   _43MB : ALIAS FOR B9[43].2;
   _43STB : ALIAS FOR B9[43].0;
   _43STPB : ALIAS FOR B9[43].1;
   _43Y : ALIAS FOR I25[2].14;
   _45_AIR_SEQ : ALIAS FOR T4[34];
   _45_AIR_SEQ1 : ALIAS FOR T4[34].PRE;
   _45_AIR_SEQ2 : ALIAS FOR T4[34].ACC;
   _45_SEQ_AIR : ALIAS FOR O12.15;
   _45AUTO : ALIAS FOR B9[45].4;
   _45HAND : ALIAS FOR B9[45].3;
   _45M : ALIAS FOR O25[8].7;
   _45MB : ALIAS FOR B9[45].2;
   _45STB : ALIAS FOR B9[45].0;
   _45STPB : ALIAS FOR B9[45].1;
   _45Y : ALIAS FOR I25[0].7;
   _46AUTO : ALIAS FOR B9[46].4;
   _46HAND : ALIAS FOR B9[46].3;
   _46M : ALIAS FOR O25[8].8;
   _46MB : ALIAS FOR B9[46].2;
   _46STB : ALIAS FOR B9[46].0;
   _46STPB : ALIAS FOR B9[46].1;
   _46Y : ALIAS FOR I25[0].8;
   _47AUTO : ALIAS FOR B9[47].4;
   _47HAND : ALIAS FOR B9[47].3;
   _47M : ALIAS FOR O25[9].10;
   _47MB : ALIAS FOR B9[47].2;
   _47STB : ALIAS FOR B9[47].0;
   _47STPB : ALIAS FOR B9[47].1;
   _47Y : ALIAS FOR I25[1].10;
   _48_CIMBRIA_HM : HOUR_METER := (MOTOR_RUNNING_INPUT_1 := 1, HR_METER_DISPLAY := 24757, MAINTENANCE_ALARM := 1);
   _48_FREQ_IN : ALIAS FOR N7[10];
   _48_FREQ_OU : ALIAS FOR N7[12];
   _48_SET_SPD : ALIAS FOR N7[11];
   _48_VFD_TO : ALIAS FOR N180[2];
   _48AUTO : ALIAS FOR B9[48].4;
   _48HAND : ALIAS FOR B9[48].3;
   _48M : ALIAS FOR O25[8].3;
   _48MAI : ALIAS FOR O25[25].2;
   _48MB : ALIAS FOR B9[48].2;
   _48STB : ALIAS FOR B9[48].0;
   _48STPB : ALIAS FOR B9[48].1;
   _48Y : ALIAS FOR I25[0].3;
   _49AUTO : ALIAS FOR B9[49].4;
   _49HAND : ALIAS FOR B9[49].3;
   _49M : ALIAS FOR O25[9].9;
   _49MB : ALIAS FOR B9[49].2;
   _49STB : ALIAS FOR B9[49].0;
   _49STPB : ALIAS FOR B9[49].1;
   _49Y : ALIAS FOR I25[1].9;
   _4_LOWER_TANK_CONVAYOR_21TO23_HM : HOUR_METER := (HR_METER_DISPLAY := 1470, NEXT_SCHDL_MAINTENANCE := 2, MAINTENANCE_ALARM := 1);
   _4_LOWER_TANK_CONVAYOR_21TO23_RUNNING : BOOL;
   _4_LS_TO_5 : ALIAS FOR I25[4].10;
   _4_LS_TO_6 : ALIAS FOR I25[4].11;
   _4_TO_BC5_S : ALIAS FOR O25[11].10;
   _4_TO_BC6_S : ALIAS FOR O25[11].11;
   _4AUTO : ALIAS FOR B9[4].4;
   _4HAND : ALIAS FOR B9[4].3;
   _4M : ALIAS FOR O25[10].1;
   _4MB : ALIAS FOR B9[4].2;
   _4STB : ALIAS FOR B9[4].0;
   _4STPB : ALIAS FOR B9[4].1;
   _4Y : ALIAS FOR I25[2].1;
   _50AUTO : ALIAS FOR B9[50].4;
   _50HAND : ALIAS FOR B9[50].3;
   _50M : ALIAS FOR O25[8].14;
   _50MB : ALIAS FOR B9[50].2;
   _50STB : ALIAS FOR B9[50].0;
   _50STPB : ALIAS FOR B9[50].1;
   _50Y : ALIAS FOR I25[0].14;
   _51_FREQ_IN : ALIAS FOR N7[13];
   _51_FREQ_OU : ALIAS FOR N7[15];
   _51_INDENT_HM : HOUR_METER := (MOTOR_RUNNING_INPUT_1 := 1, HR_METER_DISPLAY := 26515, MAINTENANCE_ALARM := 1);
   _51_SET_SPD : ALIAS FOR N7[14];
   _51_VFD_TO : ALIAS FOR N180[3];
   _51AUTO : ALIAS FOR B9[51].4;
   _51HAND : ALIAS FOR B9[51].3;
   _51M : ALIAS FOR O25[8].4;
   _51MAI : ALIAS FOR O25[25].3;
   _51MB : ALIAS FOR B9[51].2;
   _51STB : ALIAS FOR B9[51].0;
   _51STPB : ALIAS FOR B9[51].1;
   _51Y : ALIAS FOR I25[0].4;
   _52_FREQ_IN : ALIAS FOR N7[16];
   _52_FREQ_OU : ALIAS FOR N7[18];
   _52_SET_SPD : ALIAS FOR N7[17];
   _52AUTO : ALIAS FOR B9[52].4;
   _52HAND : ALIAS FOR B9[52].3;
   _52M : ALIAS FOR O25[8].6;
   _52MAI : ALIAS FOR O25[25].4;
   _52MB : ALIAS FOR B9[52].2;
   _52STB : ALIAS FOR B9[52].0;
   _52STPB : ALIAS FOR B9[52].1;
   _52Y : ALIAS FOR I25[0].6;
   _53_FREQ_IN : ALIAS FOR N7[7];
   _53_FREQ_OU : ALIAS FOR N7[9];
   _53_SET_SPD : ALIAS FOR N7[8];
   _53_VFD_TO : ALIAS FOR N180[1];
   _53AUTO : ALIAS FOR B9[53].4;
   _53HAND : ALIAS FOR B9[53].3;
   _53M : ALIAS FOR O25[8].2;
   _53MAI : ALIAS FOR O25[25].1;
   _53MB : ALIAS FOR B9[53].2;
   _53STB : ALIAS FOR B9[53].0;
   _53STPB : ALIAS FOR B9[53].1;
   _53Y : ALIAS FOR I25[0].2;
   _54AUTO : ALIAS FOR B9[54].4;
   _54HAND : ALIAS FOR B9[54].3;
   _54M : ALIAS FOR O25[11].3;
   _54MB : ALIAS FOR B9[54].2;
   _54STB : ALIAS FOR B9[54].0;
   _54STPB : ALIAS FOR B9[54].1;
   _54Y : ALIAS FOR I25[3].3;
   _55_FREQ_IN : ALIAS FOR N7[4];
   _55_FREQ_OU : ALIAS FOR N7[6];
   _55_SET_SPD : ALIAS FOR N7[5];
   _55AUTO : ALIAS FOR B9[55].4;
   _55HAND : ALIAS FOR B9[55].3;
   _55M : ALIAS FOR O25[8].1;
   _55MB : ALIAS FOR B9[55].2;
   _55STB : ALIAS FOR B9[55].0;
   _55STPB : ALIAS FOR B9[55].1;
   _55Y : ALIAS FOR I25[0].1;
   _56AUTO : ALIAS FOR B9[56].4;
   _56HAND : ALIAS FOR B9[56].3;
   _56M : ALIAS FOR O25[11].2;
   _56MB : ALIAS FOR B9[56].2;
   _56STB : ALIAS FOR B9[56].0;
   _56STPB : ALIAS FOR B9[56].1;
   _56Y : ALIAS FOR I25[3].2;
   _57AUTO : ALIAS FOR B9[57].4;
   _57HAND : ALIAS FOR B9[57].3;
   _57M : ALIAS FOR O25[9].6;
   _57MB : ALIAS FOR B9[57].2;
   _57STB : ALIAS FOR B9[57].0;
   _57STPB : ALIAS FOR B9[57].1;
   _57Y : ALIAS FOR I25[1].6;
   _5_LOWER_CROSS_BELT_HM : HOUR_METER := (HR_METER_DISPLAY := 2452, NEXT_SCHDL_MAINTENANCE := 2, MAINTENANCE_ALARM := 1);
   _5_LOWER_CROSS_BELT_RUNNING : BOOL;
   _5AUTO : ALIAS FOR B9[5].4;
   _5HAND : ALIAS FOR B9[5].3;
   _5M : ALIAS FOR O25[10].2;
   _5MB : ALIAS FOR B9[5].2;
   _5STB : ALIAS FOR B9[5].0;
   _5STPB : ALIAS FOR B9[5].1;
   _5Y : ALIAS FOR I25[2].2;
   _6AUTO : ALIAS FOR B9[6].4;
   _6HAND : ALIAS FOR B9[6].3;
   _6M : ALIAS FOR O25[10].3;
   _6MB : ALIAS FOR B9[6].2;
   _6STB : ALIAS FOR B9[6].0;
   _6STPB : ALIAS FOR B9[6].1;
   _6Y : ALIAS FOR I25[2].3;
   _700_AIR_GA : ALIAS FOR I8.3;
   _700_METER : ALIAS FOR I8.2;
   _700_PROBE : ALIAS FOR T22[9];
   _700_TREAT : ALIAS FOR I7.3;
   _700G_13_CL : ALIAS FOR B21[70].1;
   _700G_13_OP : ALIAS FOR B21[70].0;
   _700G_CLOSE : ALIAS FOR O12.9;
   _700G_OPEN : ALIAS FOR O12.8;
   _701_AIR_GA : ALIAS FOR I8.5;
   _701_FB : ALIAS FOR B21[1].3;
   _701_K_BYPA : ALIAS FOR I8.1;
   _701_K_TREA : ALIAS FOR I8.0;
   _701_METER : ALIAS FOR I8.4;
   _701_RB : ALIAS FOR B21[1].4;
   _701_REV_CN : ALIAS FOR C5[3];
   _701_STP : ALIAS FOR B21[1].2;
   _701_TRUCK_REVERSING_BELT_HM : HOUR_METER := (HR_METER_DISPLAY := 5981, NEXT_SCHDL_MAINTENANCE := 2, MAINTENANCE_ALARM := 1);
   _701_TRUCK_REVERSING_BELT_RUNNING : BOOL;
   _701F_HPB : ALIAS FOR B21[1].0;
   _701F_M : ALIAS FOR O25[10].11;
   _701F_OFF_T : ALIAS FOR T22[1];
   _701G_CLOSE : ALIAS FOR B21[71].13;
   _701G_OPEN : ALIAS FOR B21[71].12;
   _701K_GATE : ALIAS FOR B21[11].0;
   _701K_GATE1 : ALIAS FOR B21[11].1;
   _701K_GATE2 : ALIAS FOR B21[11].2;
   _701K_VALVE : ALIAS FOR O13.10;
   _701MR : ALIAS FOR O25[9].7;
   _701R_DELAY : ALIAS FOR T22[2];
   _701R_HPB : ALIAS FOR B21[1].1;
   _701Y : BOOL;
   _701YF : ALIAS FOR I25[2].11;
   _701YR : ALIAS FOR I25[1].7;
   _702_CLEAN_JUMP_BELT_HM : HOUR_METER := (HR_METER_DISPLAY := 3983, NEXT_SCHDL_MAINTENANCE := 2, MAINTENANCE_ALARM := 1);
   _702B : ALIAS FOR B21[2].2;
   _702H_START : ALIAS FOR B21[2].0;
   _702H_STOP : ALIAS FOR B21[2].1;
   _702M : ALIAS FOR O25[9].4;
   _702Y : ALIAS FOR I25[1].4;
   _703_TREATER_JUMP_BELT_HM : HOUR_METER := (HR_METER_DISPLAY := 2423, NEXT_SCHDL_MAINTENANCE := 2, MAINTENANCE_ALARM := 1);
   _703_TREATER_JUMP_BELT_RUNNING : BOOL;
   _703B : ALIAS FOR B21[3].2;
   _703H_START : ALIAS FOR B21[3].0;
   _703H_STOP : ALIAS FOR B21[3].1;
   _703M : ALIAS FOR O25[9].14;
   _703Y : ALIAS FOR I25[1].14;
   _704B : ALIAS FOR B21[4].2;
   _704H_START : ALIAS FOR B21[4].0;
   _704H_STOP : ALIAS FOR B21[4].1;
   _704M : ALIAS FOR O25[8].11;
   _704Y : ALIAS FOR I25[0].13;
   _705B : ALIAS FOR B21[5].2;
   _705H_START : ALIAS FOR B21[5].0;
   _705H_STOP : ALIAS FOR B21[5].1;
   _705M : ALIAS FOR O25[10].12;
   _705Y : ALIAS FOR I25[2].12;
   _705YA : ALIAS FOR I25[4].15;
   _706B : ALIAS FOR B21[6].2;
   _706H_START : ALIAS FOR B21[6].0;
   _706H_STOP : ALIAS FOR B21[6].1;
   _706M : ALIAS FOR O25[9].11;
   _706Y : ALIAS FOR I25[1].11;
   _707B : ALIAS FOR B21[7].2;
   _707M : ALIAS FOR O25[11].0;
   _707Y : ALIAS FOR I25[3].0;
   _708_BOT_CN : ALIAS FOR C5[5];
   _708G_BIN_1 : ALIAS FOR O9.15;
   _708G_BIN_2 : ALIAS FOR I7.4;
   _708G_CB13 : ALIAS FOR B21[8].0;
   _708G_CB131 : ALIAS FOR B21[8].1;
   _708G_CB132 : ALIAS FOR B21[8].2;
   _708G_HOLD : ALIAS FOR B21[8].3;
   _708G_HOLD1 : ALIAS FOR B21[8].6;
   _708G_RELEA : ALIAS FOR B21[8].4;
   _708G_RESET : ALIAS FOR B21[8].5;
   _709_BOT_CN : ALIAS FOR C5[6];
   _709G_BIN_1 : ALIAS FOR O10.15;
   _709G_BIN_2 : ALIAS FOR I7.5;
   _709G_CB19 : ALIAS FOR B21[9].0;
   _709G_CB191 : ALIAS FOR B21[9].1;
   _709G_CB192 : ALIAS FOR B21[9].2;
   _709G_HOLD : ALIAS FOR B21[9].3;
   _709G_HOLD1 : ALIAS FOR B21[9].6;
   _709G_RELEA : ALIAS FOR B21[9].4;
   _709G_RESET : ALIAS FOR B21[9].5;
   _709G_RUN_T : ALIAS FOR T22[8];
   _709G_TREAT : ALIAS FOR B21[9].7;
   _709G_TREAT1 : ALIAS FOR T22[10];
   _7AUTO : ALIAS FOR B9[7].4;
   _7HAND : ALIAS FOR B9[7].3;
   _7MB : ALIAS FOR B9[7].2;
   _7STB : ALIAS FOR B9[7].0;
   _7STPB : ALIAS FOR B9[7].1;
   _8AUTO : ALIAS FOR B9[8].4;
   _8HAND : ALIAS FOR B9[8].3;
   _8MB : ALIAS FOR B9[8].2;
   _8STB : ALIAS FOR B9[8].0;
   _8STPB : ALIAS FOR B9[8].1;
   _9_AIR_SV : ALIAS FOR O24[7].6;
   _9_BYPSS_GT : ALIAS FOR I24[6].1;
   _9_CAL_MOV : ALIAS FOR O24[7].2;
   _9_CAL_VALV : ALIAS FOR I24[6].5;
   _9_DRIP_GAT : ALIAS FOR O24[7].7;
   _9_GATE_SV : ALIAS FOR O24[7].0;
   _9_GATE_SV1 : ALIAS FOR O24[7].1;
   _9_SL_SW : ALIAS FOR B9[9].6;
   _9_SLW_SPEE : ALIAS FOR I25[3].12;
   _9_STP_SPEE : ALIAS FOR I25[3].13;
   _9_TREAT_MV : ALIAS FOR I24[6].6;
   _9_TREATER : ALIAS FOR I24[6].7;
   _9_TREATER_CONVAYOR_HM : HOUR_METER := (HR_METER_DISPLAY := 4578, NEXT_SCHDL_MAINTENANCE := 2, MAINTENANCE_ALARM := 1);
   _9_TREATER_CONVAYOR_RUNNING : BOOL;
   _9_TRT_M_ST : ALIAS FOR I24[6].3;
   _9_TRT_M_ST1 : ALIAS FOR I24[6].4;
   _9_TRT_MB : ALIAS FOR B3[9].0;
   _9_TRT_MOV : ALIAS FOR O24[7].4;
   _9_TRT_STB : ALIAS FOR B3[9].1;
   _9_TRT_STPB : ALIAS FOR B3[9].2;
   _9AUTO : ALIAS FOR B9[9].4;
   _9HAND : ALIAS FOR B9[9].3;
   _9M : ALIAS FOR O25[8].10;
   _9MB : ALIAS FOR B9[9].2;
   _9STB : ALIAS FOR B9[9].0;
   _9STPB : ALIAS FOR B9[9].1;
   _9Y : ALIAS FOR I25[0].10;
   _9YB : ALIAS FOR B9[9].5;
   A16 : INT[250] := ([24] := '0 ', [25] := '0 ', [26] := '0 ', [48] := '0 ', [110] := 'ge', [140] := 'ha', [150] := '10', [200] := 'cl', [210] := 'ov', [240] := 'le');
   A18 : INT[100] := ([13] := '9$00');
   A_ACC : ALIAS FOR N10[11];
   A_ACC_SEC : ALIAS FOR N10[13];
   A_HOLD_B : ALIAS FOR B3[1].4;
   A_HOLD_MB : ALIAS FOR B3[1].3;
   A_HOLD_REL : ALIAS FOR B3[1].5;
   A_MAIN_CNT : ALIAS FOR C5[0].PRE;
   A_MAIN_CNT1 : ALIAS FOR C5[0].ACC;
   A_MAIN_TRE : ALIAS FOR C5[0];
   A_PRESET : ALIAS FOR N10[10];
   A_PRESET_S : ALIAS FOR N10[12];
   A_RESET_PB : ALIAS FOR B3[1].2;
   A_SET : ALIAS FOR B3[1].6;
   A_STB_AUTO : ALIAS FOR B3[1].0;
   A_STPB_AUT : ALIAS FOR B3[1].1;
   A_TREATER : ALIAS FOR I24[6].8;
   A_TREATER1 : ALIAS FOR T4[59];
   ALARM_FIEL : ALIAS FOR T11[7];
   ALARM_HAND : ALIAS FOR B3[0].10;
   ALARM_HMI : ALIAS FOR B3[0].6;
   ALARM_HORN : ALIAS FOR O25[11].15;
   ALARM_HORN1 : ALIAS FOR O12.14;
   ALARM_INIT : ALIAS FOR B3[0].4;
   ALARM_LIGH : ALIAS FOR O13.15;
   ALARM_LT_O : ALIAS FOR T11[3];
   ALARM_SILE : ALIAS FOR I25[4].7;
   ALARM_SILE1 : ALIAS FOR I7.13;
   ALARM_SILE2 : ALIAS FOR B3[0].3;
   ALARM_SILE3 : ALIAS FOR B3[0].5;
   ALARM_SILE4 : ALIAS FOR B3[0].9;
   ALRM_LIGHT : ALIAS FOR O25[11].14;
   ALRM_SILEN : ALIAS FOR B3[0].7;
   Always_On : BOOL := 1;
   Analog : AI[160] := ([0].In := 104.0, [0].RawMin := 147.0, [0].RawMax := 16384.0, [0].EUMax := 3770.0, [1].In := 131.0, [1].RawMin := 147.0, [1].RawMax := 16384.0, [1].EUMax := 3770.0, [2].In := 1848.0, [2].RawMin := 1884.0, [2].RawMax := 16384.0, [2].EUMax := 4000.0, [20].In := 28816.0, [20].RawMin := 31000.0, [20].EUMax := 3200.0, [20].Out := 2974.5547, [21].In := 30336.0, [21].RawMax := 31000.0, [21].EUMax := 3200.0, [21].Out := 3131.458, [22].In := 30064.0, [22].RawMax := 31000.0, [22].EUMax := 3200.0, [22].Out := 3103.3806, [23].In := 7360.0, [23].RawMax := 31000.0, [23].EUMax := 3200.0, [23].Out := 759.74194, [24].In := 9136.0, [24].RawMax := 31000.0, [24].EUMax := 3200.0, [24].Out := 943.0709, [25].In := 28656.0, [25].RawMax := 31000.0, [25].EUMax := 3200.0, [25].Out := 2958.0386, [26].In := 28944.0, [26].RawMax := 31000.0, [26].EUMax := 3200.0, [26].Out := 2987.7676);
   B12 : DINT[100];
   B15 : DINT[100] := ([16] := 2#0000_0000_0000_0000_0000_0000_0000_0011, [17] := 2#0000_0000_0000_0000_0000_0000_0000_0011, [21] := 2#0000_0000_0000_0000_0000_0000_0000_0011, [22] := 2#0000_0000_0000_0000_0000_0000_0000_0011, [23] := 2#0000_0000_0000_0000_0000_0000_0000_0011, [30] := 2#0000_0000_0000_0000_0000_0000_0000_0011);
   B17 : DINT[30] := ([11] := 2#0000_0000_0000_0000_0000_0000_0000_0010, [12] := 2#0000_0000_0000_0000_0000_0000_0000_0111, [13] := 2#0000_0000_0000_0000_0000_0000_0000_0111, [14] := 2#0000_0000_0000_0000_0000_0000_0000_0010, [15] := 2#0000_0000_0000_0000_0000_0000_0000_0010, [16] := 2#0000_0000_0000_0000_0000_0000_0000_0111, [17] := 2#0000_0000_0000_0000_0000_0000_0000_0111, [21] := 2#0000_0000_0000_0000_0000_0000_0000_0010, [22] := 2#0000_0000_0000_0000_0000_0000_0000_0111, [23] := 2#0000_0000_0000_0000_0000_0000_0000_0111, [24] := 2#0000_0000_0000_0000_0000_0000_0000_0010, [25] := 2#0000_0000_0000_0000_0000_0000_0000_0111, [26] := 2#0000_0000_0000_0000_0000_0000_0000_0010);
   B183 : DINT[1] := ([0] := 2#0000_0000_0000_0000_0000_0000_0000_0001);
   B184 : DINT[1] := ([0] := 2#0000_0000_0000_0000_0000_0000_0000_0010);
   B194 : DINT[1];
   B204 : DINT[1];
   B21 : DINT[255];
   B214 : DINT[1];
   B224 : DINT[1] := ([0] := 2#0000_0000_0000_0000_0000_0000_0000_0010);
   B234 : DINT[1];
   B243 : DINT[1] := ([0] := 2#0000_0000_0000_0000_0000_0000_0000_0011);
   B244 : DINT[1] := ([0] := 2#0000_0000_0000_0000_0000_0000_0000_0010);
   B253 : DINT[100] := ([0] := 2#0000_0000_0000_0000_0000_0000_0000_0011);
   B254 : DINT[1] := ([0] := 2#0000_0000_0000_0000_0000_0000_0000_0010);
   B3 : DINT[250] := ([0] := 2#0000_0000_0000_0000_0000_0010_1011_0000, [101] := 2#0000_0000_0000_0000_0000_0000_0000_0010, [102] := 2#0000_0000_0000_0000_0000_0000_1000_0001);
   B9 : DINT[150] := ([1] := 2#0000_0000_0000_0000_0000_0000_0001_0100, [35] := 2#0000_0000_0000_0000_0000_0000_0001_0100, [42] := 2#0000_0000_0000_0000_0000_0000_0001_0100, [43] := 2#0000_0000_0000_0000_0000_0000_0011_0100, [45] := 2#0000_0000_0000_0000_0000_0000_0001_0100, [46] := 2#0000_0000_0000_0000_0000_0000_0001_0100, [48] := 2#0000_0000_0000_0000_0000_0000_0001_0100, [49] := 2#0000_0000_0000_0000_0000_0000_0001_0100, [50] := 2#0000_0000_0000_0000_0000_0000_0000_1000, [51] := 2#0000_0000_0000_0000_0000_0000_0001_0100, [52] := 2#0000_0000_0000_0000_0000_0000_0001_0100, [53] := 2#0000_0000_0000_0000_0000_0000_0001_0100, [54] := 2#0000_0000_0000_0000_0000_0000_0001_0100, [55] := 2#0000_0000_0000_0000_0000_0000_0001_0100, [57] := 2#0000_0000_0000_0000_0000_0000_0001_0100, [102] := 2#0000_0000_0000_0000_0000_0000_0000_1000, [103] := 2#0000_0000_0000_0000_0000_0000_0000_1000, [107] := 2#0000_0000_0000_0000_0000_0000_0011_0100, [108] := 2#0000_0000_0000_0000_0000_0000_0001_0100, [122] := 2#0000_0000_0000_0000_0000_0000_0001_0100, [123] := 2#0000_0000_0000_0000_0000_0000_0001_0100);
   Beta : BOOL := 1;
   BIN_1_CLOSE : BOOL;
   BIN_1_OPEN : BOOL;
   BIN_2_CLOSE : BOOL;
   BIN_2_OPEN : BOOL;
   BIN_3_CLOSE : BOOL;
   BIN_3_OPEN : BOOL;
   BIN_4_CLOSE : BOOL;
   BIN_4_OPEN : BOOL;
   BIN_5_CLOSE : BOOL;
   BIN_5_OPEN : BOOL;
   BIN_6_CLOSE : BOOL;
   BIN_6_OPEN : BOOL;
   BIN_7_CLOSE : BOOL;
   BIN_7_OPEN : BOOL;
   Bin_Config : BOOL := 1;
   C5 : COUNTER[50] := ([0].PRE := 3000, [1].ACC := 5, [1].DN := 1, [2].PRE := 3000, [3].PRE := 2, [4].PRE := 400000, [5].PRE := 5000, [5].CU := 1, [6].PRE := 9999, [6].CU := 1, [11].PRE := 1200, [12].PRE := 30, [13].PRE := 3000, [14].PRE := 36, [15].PRE := 1500, [16].PRE := 3000, [17].PRE := 3000, [21].PRE := 3000, [22].PRE := 3000, [23].PRE := 3000, [24].PRE := 3000, [25].PRE := 3000, [26].PRE := 3000, [27].CU := 1, [28].CU := 1, [29].CU := 1, [30].PRE := 20000, [32].PRE := 20000, [33].PRE := 20000, [34].PRE := 20000, [35].PRE := 20000, [36].PRE := 20000, [37].PRE := 20000, [38].PRE := 20000, [39].PRE := 20000);
   CAL_K_FACT : ALIAS FOR F8[0];
   CAL_RESET : ALIAS FOR B15[50].0;
   Calibration_Max : REAL := 4000.0;
   CG13_METR : ALIAS FOR I8.15;
   CG_13_AIR : ALIAS FOR I8.13;
   CG_19_AIR : ALIAS FOR I8.12;
   CG_19_METR : ALIAS FOR I8.14;
   CHEM_PUMP_1 : STRING := 'water';
   CHEM_PUMP_10 : STRING := 'oil';
   CHEM_PUMP_11 : STRING := 'apron';
   CHEM_PUMP_12 : STRING := 'stamina';
   CHEM_PUMP_13 : STRING := 'TEST13';
   CHEM_PUMP_14 : STRING := 'oil';
   CHEM_PUMP_15 : STRING := 'red';
   CHEM_PUMP_2 : STRING := 'alba red';
   CHEM_PUMP_3 : STRING := 'evergol';
   CHEM_PUMP_4 : STRING := 'macho';
   CHEM_PUMP_5 : STRING := 'vib ex';
   CHEM_PUMP_6 : STRING := 'bio st';
   CHEM_PUMP_7 : STRING := 'tbz';
   CHEM_PUMP_8 : STRING := 'wuxal';
   CHEM_PUMP_9 : STRING := 'BLUE';
   CIMBRA_BIN : ALIAS FOR I25[3].10;
   CIMBRIA_BI : ALIAS FOR B15[30].0;
   CIMBRIA_BI1 : ALIAS FOR B15[30].1;
   CIMBRIA_BIN_EMPTY : BOOL;
   CIMBRIA_BIN_FULL : BOOL;
   CIMBRIA_FAN_ON : BOOL := 1;
   CIMBRIA_FAN_SPD_INPUT : DINT := 30;
   CIMBRIA_HI : ALIAS FOR B15[30].2;
   CIMBRIA_OUTPUT_SPD : DINT := 30;
   Cleaning_Motors : udt_Motor[100] := ([0].Motor_Control.Motor_Amps := 1.3896561, [1].Motor_Control.Motor_Amps := 1.006918, [2].Motor_Control.Motor_Amps := 0.8792738, [3].Motor_Control.Motor_Amps := 2.5666564);
   CLR_SORT_ASP_DELAY : TIMER := (PRE := 5000, ACC := 5002, EN := 1, DN := 1);
   CLR_SORT_ASPBLR_DELAY : TIMER := (PRE := 5000, ACC := 5004, EN := 1, DN := 1);
   CLR_SORT_LEG_DELAY : TIMER := (PRE := 5000, ACC := 5003, EN := 1, DN := 1);
   CLR_SORT_LEG_SPD10 : ALIAS FOR Local:0:I.Data.3;
   CLR_SORT_LEG_SPD20 : ALIAS FOR Local:0:I.Data.4;
   CONC13_COL : ALIAS FOR N7[93];
   CONC13_OP : ALIAS FOR A18[3];
   CONC13_PUM : ALIAS FOR N7[83];
   CONC13_SET : ALIAS FOR A18[0];
   CONC13_SET1 : ALIAS FOR B21[8].14;
   CONC19_COL : ALIAS FOR N7[99];
   CONC19_OP : ALIAS FOR A18[13];
   CONC19_PUM : ALIAS FOR N7[89];
   CONC19_SET : ALIAS FOR B21[9].14;
   CONC_13_NO : ALIAS FOR B21[8].15;
   CONC_19_NO : ALIAS FOR B21[9].15;
   CONC_19_SE : ALIAS FOR A18[10];
   ConcretePlantIn : DINT := 2;
   ConcretePlantOut : DINT := 1; {produced}
   Config_Save_Binss : BOOL;
   ConfigureVariety : Variety;
   Consumed : DINT;
   CP_Remote_Air_Gate_On : DINT; {produced}
   CP_Remote_Air_Gate_Open_In : DINT;
   CP_Remote_Andco_Auto_In : DINT;
   CP_Remote_Andoc_Out : udt_Andco_Remote_Out[32]; {produced}
   CP_Remote_Belt_In : udt_Motor_Remote_In[10] := ([1].Spd_10_Out := 1, [1].Amps := -0.32500002, [2].Spd_10_Out := 1, [2].Amps := -0.425, [3].Spd_10_Out := 1, [3].Amps := -0.5125);
   CP_Remote_Belt_Start : DINT; {produced}
   CP_Remote_Leg_In : udt_Motor_Remote_In := (Spd_20_Out := 1, Spd_10_Out := 1, Amps := -0.22500001);
   CP_Remote_Leg_Start : DINT; {produced}
   cpBinGateRates : DINT[50] := ([1] := 73, [3] := 180, [5] := 531, [7] := 117, [10] := 147, [13] := 269, [19] := 173);
   cpBINOPEN : DINT;
   cpCleanBulk : BOOL;
   cpTicketBinActive : DINT;
   cpTicketBinSet : DINT;
   cpVAR_BINARRAY : STRING[50] := ([1] := '823019-Diva Spring-Certified-WSU -SWW Seed Wheat', [3] := '823007-WB 6121 spring-Certified - Monsanto  - SWW Seed Wheat', [4] := 'reg duet', [5] := '823001-ArtDeco-Certified-Limagrain -SWW Seed Wheat', [10] := '823007-WB 6121 spring-Certified-Monsanto -SWW Seed Wheat', [11] := '823014-Skiles-Certified-OSU -SWW Seed Wheat', [20] := '823010-Bobtail-Certified-OSU -SWW Seed Wheat');
   cpVAR_CNT_ONS : DINT;
   cpVarTrimTemp : STRING := '823026';
   Dev : DINT := 6145; {produced}
   DIST_MOVE : ALIAS FOR I3.10;
   DIST_TO_CL : ALIAS FOR I7.2;
   DS_CLEAN_B : ALIAS FOR O13.5;
   DS_DLY_OFF : ALIAS FOR T4[33];
   DS_M : ALIAS FOR O24[1].0;
   DS_M_B : ALIAS FOR B3[101].0;
   DS_MOV_CCW : ALIAS FOR B3[100].13;
   DS_MOV_CW : ALIAS FOR B3[100].12;
   DS_MOVE_SE : ALIAS FOR T4[32];
   DS_POS8 : ALIAS FOR O13.7;
   DS_POS9 : ALIAS FOR O13.8;
   DS_POS_1 : ALIAS FOR I24[0].2;
   DS_POS_10 : ALIAS FOR I24[0].11;
   DS_POS_11 : ALIAS FOR B3[100].11;
   DS_POS_1_B : ALIAS FOR B3[100].2;
   DS_POS_2 : ALIAS FOR I24[0].3;
   DS_POS_2_B : ALIAS FOR B3[100].3;
   DS_POS_3 : ALIAS FOR I24[0].4;
   DS_POS_3_B : ALIAS FOR B3[100].4;
   DS_POS_4 : ALIAS FOR I24[0].5;
   DS_POS_4_B : ALIAS FOR B3[100].5;
   DS_POS_5 : ALIAS FOR I24[0].6;
   DS_POS_5_B : ALIAS FOR B3[100].6;
   DS_POS_6 : ALIAS FOR I24[0].7;
   DS_POS_6_B : ALIAS FOR B3[100].7;
   DS_POS_7 : ALIAS FOR I24[0].8;
   DS_POS_7_B : ALIAS FOR B3[100].8;
   DS_POS_8 : ALIAS FOR I24[0].9;
   DS_POS_8_B : ALIAS FOR B3[100].9;
   DS_POS_9 : ALIAS FOR I24[0].10;
   DS_POS_9_B : ALIAS FOR B3[100].10;
   DS_SEEK_1 : ALIAS FOR B3[102].1;
   DS_SEEK_10 : ALIAS FOR B3[102].10;
   DS_SEEK_2 : ALIAS FOR B3[102].2;
   DS_SEEK_3 : ALIAS FOR B3[102].3;
   DS_SEEK_4 : ALIAS FOR B3[102].4;
   DS_SEEK_5 : ALIAS FOR B3[102].5;
   DS_SEEK_6 : ALIAS FOR B3[102].6;
   DS_SEEK_7 : ALIAS FOR B3[102].7;
   DS_SEEK_8 : ALIAS FOR B3[102].8;
   DS_SEEK_9 : ALIAS FOR B3[102].9;
   DS_SET_IN : ALIAS FOR N10[0];
   DS_SP_UP_B : ALIAS FOR B3[100].0;
   DS_SPOUT_C : ALIAS FOR O24[1].3;
   DS_SPOUT_C1 : ALIAS FOR O24[1].4;
   DS_SPOUT_C2 : ALIAS FOR B3[101].3;
   DS_SPOUT_C3 : ALIAS FOR B3[101].4;
   DS_SPOUT_D : ALIAS FOR I24[0].1;
   DS_SPOUT_D1 : ALIAS FOR O24[1].1;
   DS_SPOUT_D2 : ALIAS FOR B3[100].1;
   DS_SPOUT_D3 : ALIAS FOR B3[101].1;
   DS_SPOUT_U : ALIAS FOR I24[0].0;
   DS_SPOUT_U1 : ALIAS FOR O24[1].2;
   DS_SPOUT_U2 : ALIAS FOR B3[101].2;
   DS_START_M : ALIAS FOR B3[102].11;
   DS_STOP_MO : ALIAS FOR B3[102].0;
   DS_T21 : ALIAS FOR O13.0;
   DS_T22 : ALIAS FOR O13.1;
   DS_T23 : ALIAS FOR O13.9;
   DS_T231 : ALIAS FOR O13.2;
   DS_T24 : ALIAS FOR O13.3;
   DS_T25 : ALIAS FOR O13.4;
   DS_T26 : ALIAS FOR O13.6;
   F8 : REAL[27] := ([0] := 1.2, [1] := 1.0, [2] := 14748.0, [3] := 1.0, [4] := 15440.0, [5] := 1.0, [6] := 14244.0, [7] := 1.0, [8] := 13454.0, [9] := 1.0, [10] := 14460.0, [11] := 1.0, [12] := 6343.0, [13] := 1.0, [14] := 8758.0, [15] := 1.0, [16] := 15944.0, [17] := 1.0, [18] := 15184.0, [19] := 1.0, [20] := 15741.0, [21] := 1.0, [22] := 15276.0, [23] := 1.0, [24] := 14611.0, [25] := 1.0, [26] := 15145.0);
   Gates : STRING;
   hCLR_SORT_LEG_SPD10 : BOOL := 1;
   hCLR_SORT_LEG_SPD20 : BOOL := 1;
   hCLR_SORT_STB : BOOL;
   hCLR_SORT_STRT : BOOL;
   hN_RECVING_PIT_GATE_CLSPB : BOOL;
   hN_RECVING_PIT_GATE_OPNPB : BOOL;
   hSURGE_BIN_HI : BOOL;
   hSURGE_BIN_LO : BOOL;
   I1 : ALIAS FOR R1S0_AENTR:1:I.Data;
   I16 : INT[16] := ([0] := 2#0011_1001_1001_1100, [1] := 2#0011_1100_0101_0000, [2] := 2#0011_0111_1010_0100, [3] := 2#0011_0100_1000_1110, [4] := 2#0011_1000_0111_1100, [5] := 2#0001_1000_1100_0111, [6] := 2#0010_0010_0011_0110, [7] := 2#0011_1110_0100_1000, [8] := 2#0000_1000_0101_1010, [9] := 2#0000_1000_0101_1010, [10] := 2#0000_1000_0101_1010, [11] := 2#0000_1000_0101_1010, [12] := 2#0000_1000_0101_1010, [13] := 2#0000_1000_0101_1010, [14] := 2#0000_1000_0101_1010, [15] := 2#0000_1000_0101_1010);
   I16_0 : ALIAS FOR N20[0];
   I16_000 : ALIAS FOR I16[0];
   I16_001 : ALIAS FOR I16[1];
   I16_002 : ALIAS FOR I16[2];
   I16_003 : ALIAS FOR I16[3];
   I16_004 : ALIAS FOR I16[4];
   I16_005 : ALIAS FOR I16[5];
   I16_006 : ALIAS FOR I16[6];
   I16_007 : ALIAS FOR I16[7];
   I16_1 : ALIAS FOR N20[1];
   I16_2 : ALIAS FOR N20[2];
   I16_3 : ALIAS FOR N20[3];
   I16_4 : ALIAS FOR N20[4];
   I16_5 : ALIAS FOR N20[5];
   I16_6 : ALIAS FOR N20[6];
   I16_7 : ALIAS FOR N20[7];
   I17 : INT[16] := ([0] := 2#0011_1011_0101_0000, [1] := 2#0011_1101_0111_1101, [2] := 2#0011_1011_1010_1111, [3] := 2#0011_1001_0001_0011, [4] := 2#0011_1011_0010_1001, [5] := 2#0001_1100_1010_0101, [6] := 2#0001_1100_1010_1111, [7] := 2#0001_1100_1010_0010, [8] := 2#0000_1000_0101_1010, [9] := 2#0000_1000_0101_1010, [10] := 2#0000_1000_0101_1010, [11] := 2#0000_1000_0101_1010, [12] := 2#0000_1000_0101_1010, [13] := 2#0000_1000_0101_1010, [14] := 2#0000_1000_0101_1010, [15] := 2#0000_1000_0101_1010);
   I17_000 : ALIAS FOR I17[0];
   I17_001 : ALIAS FOR I17[1];
   I17_002 : ALIAS FOR I17[2];
   I17_003 : ALIAS FOR I17[3];
   I17_004 : ALIAS FOR I17[4];
   I17_005 : ALIAS FOR I17[5];
   I17_006 : ALIAS FOR I17[6];
   I17_007 : ALIAS FOR I17[7];
   I18 : INT[16] := ([0] := 2#0000_0101_0101_0011, [1] := 2#0000_0111_0011_1000, [2] := 2#0000_0000_1000_0011, [3] := 2#0000_0000_0110_1000, [4] := 2#0000_0111_0111_1100, [5] := 2#0000_0111_0110_0101, [6] := 2#0000_1100_1100_1101, [7] := 2#0000_1100_1100_1101, [8] := 2#0000_1000_0101_1010, [9] := 2#0000_1000_0101_1010, [10] := 2#0000_1000_0101_1010, [11] := 2#0000_1000_0101_1010, [12] := 2#0000_1000_0101_1010, [13] := 2#0000_1000_0101_1010, [14] := 2#0001_1010_1001_1101, [15] := 2#0001_1010_1001_1101);
   I18_000 : ALIAS FOR I18[0];
   I18_001 : ALIAS FOR I18[1];
   I18_002 : ALIAS FOR I18[2];
   I18_003 : ALIAS FOR I18[3];
   I18_007 : ALIAS FOR I18[7];
   I1_000_Bit00 : ALIAS FOR I1.0;
   I1_000_Bit01 : ALIAS FOR I1.1;
   I1_000_Bit02 : ALIAS FOR I1.2;
   I1_000_Bit03 : ALIAS FOR I1.3;
   I1_000_Bit04 : ALIAS FOR I1.4;
   I1_000_Bit05 : ALIAS FOR I1.5;
   I1_000_Bit06 : ALIAS FOR I1.6;
   I1_000_Bit07 : ALIAS FOR I1.7;
   I1_000_Bit08 : ALIAS FOR I1.8;
   I1_000_Bit09 : ALIAS FOR I1.9;
   I1_000_Bit10 : ALIAS FOR I1.10;
   I1_000_Bit11 : ALIAS FOR I1.11;
   I1_000_Bit12 : ALIAS FOR I1.12;
   I1_000_Bit13 : ALIAS FOR I1.13;
   I1_000_Bit14 : ALIAS FOR I1.14;
   I1_000_Bit15 : ALIAS FOR I1.15;
   I2 : ALIAS FOR R1S0_AENTR:2:I.Data;
   I24 : INT[32] := ([0] := 2#0000_0001_0000_0010, [6] := 2#0010_0000_1000_0110, [7] := 2#0010_0000_1000_0110);
   I24_000_Bit00 : ALIAS FOR I24[0].0;
   I24_000_Bit01 : ALIAS FOR I24[0].1;
   I24_000_Bit02 : ALIAS FOR I24[0].2;
   I24_000_Bit03 : ALIAS FOR I24[0].3;
   I24_000_Bit04 : ALIAS FOR I24[0].4;
   I24_000_Bit05 : ALIAS FOR I24[0].5;
   I24_000_Bit06 : ALIAS FOR I24[0].6;
   I24_000_Bit07 : ALIAS FOR I24[0].7;
   I24_000_Bit08 : ALIAS FOR I24[0].8;
   I24_000_Bit09 : ALIAS FOR I24[0].9;
   I24_000_Bit10 : ALIAS FOR I24[0].10;
   I24_000_Bit11 : ALIAS FOR I24[0].11;
   I24_004_Bit00 : ALIAS FOR I24[4].0;
   I24_004_Bit01 : ALIAS FOR I24[4].1;
   I24_004_Bit02 : ALIAS FOR I24[4].2;
   I24_004_Bit03 : ALIAS FOR I24[4].3;
   I24_004_Bit04 : ALIAS FOR I24[4].4;
   I24_004_Bit05 : ALIAS FOR I24[4].5;
   I24_004_Bit06 : ALIAS FOR I24[4].6;
   I24_004_Bit07 : ALIAS FOR I24[4].7;
   I24_004_Bit08 : ALIAS FOR I24[4].8;
   I24_004_Bit09 : ALIAS FOR I24[4].9;
   I24_004_Bit10 : ALIAS FOR I24[4].10;
   I24_004_Bit11 : ALIAS FOR I24[4].11;
   I24_004_Bit12 : ALIAS FOR I24[4].12;
   I24_006_Bit01 : ALIAS FOR I24[6].1;
   I24_006_Bit02 : ALIAS FOR I24[6].2;
   I24_006_Bit07 : ALIAS FOR I24[6].7;
   I24_006_Bit08 : ALIAS FOR I24[6].8;
   I24_006_Bit13 : ALIAS FOR I24[6].13;
   I24_021_Bit00 : ALIAS FOR I24[21].0;
   I24_021_Bit01 : ALIAS FOR I24[21].1;
   I24_021_Bit02 : ALIAS FOR I24[21].2;
   I24_021_Bit03 : ALIAS FOR I24[21].3;
   I24_021_Bit04 : ALIAS FOR I24[21].4;
   I24_021_Bit05 : ALIAS FOR I24[21].5;
   I24_021_Bit06 : ALIAS FOR I24[21].6;
   I24_021_Bit07 : ALIAS FOR I24[21].7;
   I24_021_Bit08 : ALIAS FOR I24[21].8;
   I25 : INT[32] := ([0] := 2#0101_0011_1101_1110, [1] := 2#0011_0011_0100_0010, [2] := 2#1110_0000_0100_0000, [3] := 2#1101_0000_0000_1010, [4] := 2#0110_0000_0000_1101);
   I25_000_Bit00 : ALIAS FOR I25[0].0;
   I25_000_Bit01 : ALIAS FOR I25[0].1;
   I25_000_Bit02 : ALIAS FOR I25[0].2;
   I25_000_Bit03 : ALIAS FOR I25[0].3;
   I25_000_Bit04 : ALIAS FOR I25[0].4;
   I25_000_Bit06 : ALIAS FOR I25[0].6;
   I25_000_Bit07 : ALIAS FOR I25[0].7;
   I25_000_Bit08 : ALIAS FOR I25[0].8;
   I25_000_Bit09 : ALIAS FOR I25[0].9;
   I25_000_Bit10 : ALIAS FOR I25[0].10;
   I25_000_Bit12 : ALIAS FOR I25[0].12;
   I25_000_Bit13 : ALIAS FOR I25[0].13;
   I25_000_Bit14 : ALIAS FOR I25[0].14;
   I25_000_Bit15 : ALIAS FOR I25[0].15;
   I25_001_Bit00 : ALIAS FOR I25[1].0;
   I25_001_Bit01 : ALIAS FOR I25[1].1;
   I25_001_Bit02 : ALIAS FOR I25[1].2;
   I25_001_Bit03 : ALIAS FOR I25[1].3;
   I25_001_Bit04 : ALIAS FOR I25[1].4;
   I25_001_Bit05 : ALIAS FOR I25[1].5;
   I25_001_Bit06 : ALIAS FOR I25[1].6;
   I25_001_Bit07 : ALIAS FOR I25[1].7;
   I25_001_Bit08 : ALIAS FOR I25[1].8;
   I25_001_Bit09 : ALIAS FOR I25[1].9;
   I25_001_Bit10 : ALIAS FOR I25[1].10;
   I25_001_Bit11 : ALIAS FOR I25[1].11;
   I25_001_Bit12 : ALIAS FOR I25[1].12;
   I25_001_Bit13 : ALIAS FOR I25[1].13;
   I25_001_Bit14 : ALIAS FOR I25[1].14;
   I25_001_Bit15 : ALIAS FOR I25[1].15;
   I25_002_Bit00 : ALIAS FOR I25[2].0;
   I25_002_Bit01 : ALIAS FOR I25[2].1;
   I25_002_Bit02 : ALIAS FOR I25[2].2;
   I25_002_Bit03 : ALIAS FOR I25[2].3;
   I25_002_Bit04 : ALIAS FOR I25[2].4;
   I25_002_Bit05 : ALIAS FOR I25[2].5;
   I25_002_Bit06 : ALIAS FOR I25[2].6;
   I25_002_Bit08 : ALIAS FOR I25[2].8;
   I25_002_Bit09 : ALIAS FOR I25[2].9;
   I25_002_Bit10 : ALIAS FOR I25[2].10;
   I25_002_Bit11 : ALIAS FOR I25[2].11;
   I25_002_Bit12 : ALIAS FOR I25[2].12;
   I25_002_Bit13 : ALIAS FOR I25[2].13;
   I25_002_Bit14 : ALIAS FOR I25[2].14;
   I25_002_Bit15 : ALIAS FOR I25[2].15;
   I25_003_Bit00 : ALIAS FOR I25[3].0;
   I25_003_Bit01 : ALIAS FOR I25[3].1;
   I25_003_Bit03 : ALIAS FOR I25[3].3;
   I25_003_Bit10 : ALIAS FOR I25[3].10;
   I25_003_Bit12 : ALIAS FOR I25[3].12;
   I25_003_Bit13 : ALIAS FOR I25[3].13;
   I25_003_Bit14 : ALIAS FOR I25[3].14;
   I25_003_Bit15 : ALIAS FOR I25[3].15;
   I25_004_Bit00 : ALIAS FOR I25[4].0;
   I25_004_Bit01 : ALIAS FOR I25[4].1;
   I25_004_Bit02 : ALIAS FOR I25[4].2;
   I25_004_Bit03 : ALIAS FOR I25[4].3;
   I25_004_Bit06 : ALIAS FOR I25[4].6;
   I25_004_Bit07 : ALIAS FOR I25[4].7;
   I25_004_Bit14 : ALIAS FOR I25[4].14;
   I2_000_Bit00 : ALIAS FOR I2.0;
   I2_000_Bit02 : ALIAS FOR I2.2;
   I2_000_Bit03 : ALIAS FOR I2.3;
   I2_000_Bit05 : ALIAS FOR I2.5;
   I2_000_Bit06 : ALIAS FOR I2.6;
   I2_000_Bit07 : ALIAS FOR I2.7;
   I2_000_Bit08 : ALIAS FOR I2.8;
   I2_000_Bit09 : ALIAS FOR I2.9;
   I2_000_Bit10 : ALIAS FOR I2.10;
   I2_000_Bit11 : ALIAS FOR I2.11;
   I2_000_Bit12 : ALIAS FOR I2.12;
   I2_000_Bit13 : ALIAS FOR I2.13;
   I2_000_Bit14 : ALIAS FOR I2.14;
   I3 : ALIAS FOR R1S0_AENTR:3:I.Data;
   I3_000_Bit00 : ALIAS FOR I3.0;
   I3_000_Bit01 : ALIAS FOR I3.1;
   I3_000_Bit02 : ALIAS FOR I3.2;
   I3_000_Bit03 : ALIAS FOR I3.3;
   I3_000_Bit04 : ALIAS FOR I3.4;
   I3_000_Bit05 : ALIAS FOR I3.5;
   I3_000_Bit06 : ALIAS FOR I3.6;
   I3_000_Bit07 : ALIAS FOR I3.7;
   I3_000_Bit08 : ALIAS FOR I3.8;
   I3_000_Bit09 : ALIAS FOR I3.9;
   I3_000_Bit10 : ALIAS FOR I3.10;
   I3_000_Bit11 : ALIAS FOR I3.11;
   I3_000_Bit12 : ALIAS FOR I3.12;
   I3_000_Bit14 : ALIAS FOR I3.14;
   I4 : ALIAS FOR R1S0_AENTR:4:I.Data;
   I4_000_Bit00 : ALIAS FOR I4.0;
   I4_000_Bit02 : ALIAS FOR I4.2;
   I4_000_Bit04 : ALIAS FOR I4.4;
   I4_000_Bit09 : ALIAS FOR I4.9;
   I4_000_Bit10 : ALIAS FOR I4.10;
   I4_000_Bit11 : ALIAS FOR I4.11;
   I4_000_Bit12 : ALIAS FOR I4.12;
   I4_000_Bit13 : ALIAS FOR I4.13;
   I4_000_Bit14 : ALIAS FOR I4.14;
   I4_000_Bit15 : ALIAS FOR I4.15;
   I5 : ALIAS FOR R1S0_AENTR:5:I.Data;
   I6 : ALIAS FOR R1S0_AENTR:6:I.Data;
   I7 : ALIAS FOR R1S0_AENTR:7:I.Data;
   I7_000_Bit02 : ALIAS FOR I7.2;
   I7_000_Bit03 : ALIAS FOR I7.3;
   I7_000_Bit04 : ALIAS FOR I7.4;
   I7_000_Bit05 : ALIAS FOR I7.5;
   I7_000_Bit13 : ALIAS FOR I7.13;
   I7_000_Bit14 : ALIAS FOR I7.14;
   I7_000_Bit15 : ALIAS FOR I7.15;
   I8 : ALIAS FOR R1S0_AENTR:8:I.Data;
   I8_000_Bit00 : ALIAS FOR I8.0;
   I8_000_Bit02 : ALIAS FOR I8.2;
   I8_000_Bit03 : ALIAS FOR I8.3;
   I8_000_Bit04 : ALIAS FOR I8.4;
   I8_000_Bit05 : ALIAS FOR I8.5;
   I8_000_Bit06 : ALIAS FOR I8.6;
   I8_000_Bit07 : ALIAS FOR I8.7;
   I8_000_Bit08 : ALIAS FOR I8.8;
   I8_000_Bit09 : ALIAS FOR I8.9;
   I8_000_Bit10 : ALIAS FOR I8.10;
   I8_000_Bit11 : ALIAS FOR I8.11;
   I8_000_Bit12 : ALIAS FOR I8.12;
   IE8_BTR_FL : ALIAS FOR N23[0];
   indexTbl : DINT;
   indexTblOld : DINT;
   indexTRTTbl : DINT;
   InEUMax : REAL;
   K_FACTOR : ALIAS FOR N14[80];
   M0_24 : INT[3300] := ([100] := -32640, [200] := -32768, [300] := 128, [400] := -32768, [500] := -32640, [700] := -32640, [800] := -32768, [900] := -32640);
   M0_25 : INT[3300] := ([100] := -32640, [300] := -32640, [500] := 128, [600] := -32768);
   M1_24 : INT[3300];
   M1_25 : INT[3300];
   M701_SLOW : ALIAS FOR I8.6;
   M701_STOP : ALIAS FOR I8.7;
   M702_SLOW : ALIAS FOR I8.8;
   M702_STOP : ALIAS FOR I8.9;
   M703_SLOW : ALIAS FOR I8.10;
   M703_STOP : ALIAS FOR I8.11;
   MAIN_TIMER : ALIAS FOR T11[0];
   MAIN_TIMER1 : ALIAS FOR T11[1];
   MASTER_FAU : ALIAS FOR B3[0].1;
   MASTER_STO : ALIAS FOR B3[0].2;
   MTR_125_RUNNING : ALIAS FOR Local:0:I.Data.11;
   MTR_125MB : ALIAS FOR Local:5:O.Data.0;
   MTR_126_RUNNING : ALIAS FOR Local:0:I.Data.6;
   MTR_126M : ALIAS FOR Local:5:O.Data.1;
   MTR_126MB : BOOL := 1;
   MTR_127_RUNNING : ALIAS FOR Local:0:I.Data.7;
   MTR_127M : ALIAS FOR Local:5:O.Data.2;
   MTR_127MB : BOOL := 1;
   MTR_128_RUNNING : ALIAS FOR Local:0:I.Data.5;
   MTR_128M : ALIAS FOR Local:5:O.Data.3;
   MTR_128MB : BOOL := 1;
   N10 : DINT[30] := ([0] := 7, [1] := 7, [10] := 500, [12] := 3000);
   N13 : DINT[100] := ([4] := 80, [14] := 43, [24] := 35, [34] := 30, [44] := 29, [54] := 30, [64] := 30, [74] := 40, [84] := 22);
   N14 : DINT[84] := ([11] := 3173, [12] := 3523, [13] := 2924, [14] := 3485, [15] := 3442, [16] := 1402, [17] := 2895, [21] := 3209, [22] := 3053, [23] := 3621, [24] := 3332, [25] := 4010, [26] := 3739, [31] := 1, [32] := 7589, [33] := 7589, [34] := 1, [35] := 9417, [36] := 9417, [37] := 1, [38] := 10027, [39] := 10027, [40] := 1, [41] := 8, [43] := 1, [44] := 8771, [45] := 8771, [46] := 1, [47] := 8060, [48] := 8060, [49] := 1, [50] := 6101, [51] := 6101, [52] := 1, [53] := 15066, [54] := 15066, [55] := 1, [56] := 10230, [57] := 10230, [58] := 1, [59] := 9011, [60] := 9011, [61] := 1, [62] := 9440, [63] := 9440, [64] := 1, [65] := 7454, [66] := 7454, [67] := 1, [68] := 9863, [69] := 9863, [80] := 120);
   N180 : DINT[68] := ([0] := 160, [1] := 14932, [2] := 27374, [3] := 14300, [4] := 23411, [5] := 12, [7] := 3026, [8] := 239, [10] := -256, [50] := 128, [51] := 9, [52] := 220, [54] := 1, [55] := 220, [60] := 25600, [61] := 9, [62] := 220, [64] := 1024, [66] := 220);
   N181 : DINT[1];
   N182 : DINT[2] := ([0] := -9, [1] := -9);
   N190 : DINT[68] := ([0] := 14, [10] := 23340, [14] := 15, [15] := 3840, [50] := -32640, [51] := 1, [52] := 210, [54] := 14, [55] := 210, [61] := 1, [62] := 210, [64] := 25600, [65] := 14, [66] := 210);
   N191 : DINT[1];
   N192 : DINT[2] := ([0] := -9, [1] := -9);
   N193 : DINT[1] := ([0] := 9);
   N20 : DINT[30] := ([0] := 2138, [1] := 2138, [2] := 2138, [3] := 2138, [4] := 2138, [5] := 2138, [6] := 2138, [7] := 2138, [10] := 2138, [11] := 2138, [12] := 2138, [13] := 2138, [14] := 2138, [15] := 2138, [16] := 2138, [17] := 2138, [20] := 2138, [21] := 2138, [22] := 2138, [23] := 2138, [24] := 2138, [25] := 2138, [26] := 2717, [27] := 2717);
   N200 : DINT[68] := ([10] := 400, [11] := 24800, [12] := 27383, [13] := 23767, [14] := 15, [15] := 3840, [50] := -32640, [51] := 1, [52] := 200, [54] := 14, [55] := 200, [61] := 1, [62] := 200, [64] := 25600, [65] := 14, [66] := 200);
   N201 : DINT[1];
   N202 : DINT[2] := ([0] := -9, [1] := -9);
   N203 : DINT[1] := ([0] := 9);
   N210 : DINT[68] := ([0] := 14, [10] := 7040, [11] := 2, [14] := 15, [15] := 3840, [50] := -32640, [51] := 1, [52] := 240, [54] := 14, [55] := 240, [60] := 1024, [62] := 240, [64] := 25600, [65] := 14, [66] := 240);
   N211 : DINT[1];
   N212 : DINT[2] := ([0] := -9, [1] := -9);
   N213 : DINT[1] := ([0] := 9);
   N220 : DINT[68] := ([10] := 9280, [11] := 9600, [12] := 9600, [13] := 12800, [14] := 15, [15] := 3840, [50] := -32640, [51] := 1, [52] := 230, [54] := 14, [55] := 230, [61] := 1, [62] := 230, [64] := 1024, [66] := 230);
   N221 : DINT[1];
   N222 : DINT[2] := ([0] := -9, [1] := -9);
   N223 : DINT[1] := ([0] := 3);
   N23 : DINT[5] := ([0] := 11, [1] := 60, [2] := 11, [3] := 60);
   N230 : DINT[68] := ([10] := 24720, [11] := 13760, [12] := 11200, [13] := 9600, [14] := 15, [15] := 3840, [50] := -32640, [51] := 1, [52] := 220, [54] := 14, [55] := 220, [61] := 1, [62] := 220, [64] := 25600, [65] := 14, [66] := 220);
   N231 : DINT[1];
   N232 : DINT[2] := ([0] := -9, [1] := -9);